(* Logix 5000 project; controller Almacen_2 vendor 1 type 14 code 235 rev 36.11; software revision 36.00; part 2 of 2 *)
(* tags used below, declared in another part *)
   Contador_Salida_Conveyor : COUNTER;
   End_Conveyor_Rutine : BOOL;
   PosDer_Alm_5_C : BOOL;
   PosDer_Alm_5_E : BOOL;
   PosIzq_Alm_7_C : BOOL;
   PosIzq_Conv_7_C : BOOL;
   PosIzq_Conv_8_C : BOOL;
   Recuperar_Pieza : BOOL;
   Recuperar_Pieza_Desde_RutinaConveyor : BOOL;
   Reset_RutinaFinal : BOOL;
   Start_Conveyor : BOOL;
   Start_Rutine_Conveyor_2 : BOOL;
   Stop_Conveyor_2 : BOOL;
   tag_switch : BOOL;
   tag_switch2 : BOOL;
   tag_switch3 : BOOL;
   Tag_switch4 : BOOL;
   tag_switch5 : BOOL;
   tag_switch6 : BOOL;
   tag_switch7 : BOOL;
   tag_switch8 : BOOL;
   tag_switch_almacen10 : BOOL;
   tag_switch_almacen11 : BOOL;
   tag_switch_almacen12 : BOOL;
   tag_switch_almacen13 : BOOL;
   tag_switch_almacen14 : BOOL;
   tag_switch_almacen15 : BOOL;
   tag_switch_almacen16 : BOOL;
   tag_switch_almacen17 : BOOL;
   tag_switch_almacen_abrir_gripper2 : BOOL;
   tag_switch_almacen_cerrar_gripper2 : BOOL;
   tag_timer_piston : BOOL;
   tag_timer_piston2 : BOOL;
   Timer10_Recuperar_Pieza : TIMER;
   Timer11_Posicion_Recuperar_Pieza : TIMER;
   Timer1_Cambio_Direccion_CNC : TIMER;
   Timer2 : TIMER;
   Timer3_Piston_Marcadora_OFF : TIMER;
   Timer4_Piston_Camara_ON : TIMER;
   Timer5_Piston_Camara_OFF : TIMER;
   Timer6_Cambio_Direccion_Almacen : TIMER;
   Timer7_Sensor_Entrada_Salida : TIMER;
   Timer8_End_RutinaConveyor : TIMER;
   Timer9_Piston_Salida : TIMER;
   Timer_Almacen_Abrir_Gripper2 : TIMER;
   Timer_Almacen_Cerrar_Gripper2 : TIMER;
   Timer_Almacen_Entrar_Posicion1_Regreso : TIMER;
   Timer_Almacen_Posicion_1_Regreso : TIMER;
   Timer_Almacen_Posicion_Above_Conveyor3 : TIMER;
   Timer_Almacen_Posicion_Above_Conveyor4 : TIMER;
   Timer_Almacen_Posicion_Conveyor2 : TIMER;
   Timer_Almacen_Posicion_Home3 : TIMER;
   Timer_Almacen_Posicion_Home4 : TIMER;
   Timer_Almacen_Salir_Posicion1_Regreso : TIMER;
   Estops_Ok : BOOL;
   Interlocks_Ok : BOOL;
   LigthCurtain2_Ok : BOOL;
   Run_Program_Almacen2 : BOOL;
   Safety_FromTEC81 : Safety;
   Sfty_OK : BOOL;
   Start_Almacen2 : BOOL;
   Start_Conveyor_2_From_RutinaFinal : BOOL;
   Start_Motor_Alm_2 : BOOL;
   Start_RutinaFinal : BOOL;
   tag_switch_almacen1 : BOOL;
   tag_switch_almacen2 : BOOL;
   tag_switch_almacen3 : BOOL;
   tag_switch_almacen4 : BOOL;
   tag_switch_almacen5 : BOOL;
   tag_switch_almacen6 : BOOL;
   tag_switch_almacen7 : BOOL;
   tag_switch_almacen8 : BOOL;
   tag_switch_almacen9 : BOOL;
   tag_switch_almacen_abrir_gripper : BOOL;
   tag_switch_almacen_cerrar_gripper : BOOL;
   Timer_Almacen_Abrir_Gripper : TIMER;
   Timer_Almacen_Cerrar_Gripper : TIMER;
   Timer_Almacen_Entrar_Posicion1 : TIMER;
   Timer_Almacen_Posicion1 : TIMER;
   Timer_Almacen_Posicion_Above_Conveyor : TIMER;
   Timer_Almacen_Posicion_Above_Conveyor2 : TIMER;
   Timer_Almacen_Posicion_Conveyor : TIMER;
   Timer_Almacen_Posicion_Giro_A_Conveyor : TIMER;
   Timer_Almacen_Posicion_Home : TIMER;
   Timer_Almacen_Posicion_Home2 : TIMER;
   Timer_Almacen_Salir_Posicion1 : TIMER;
(* MainProgram, continued *)

ROUTINE RutinaConveyor   (* ladder *)
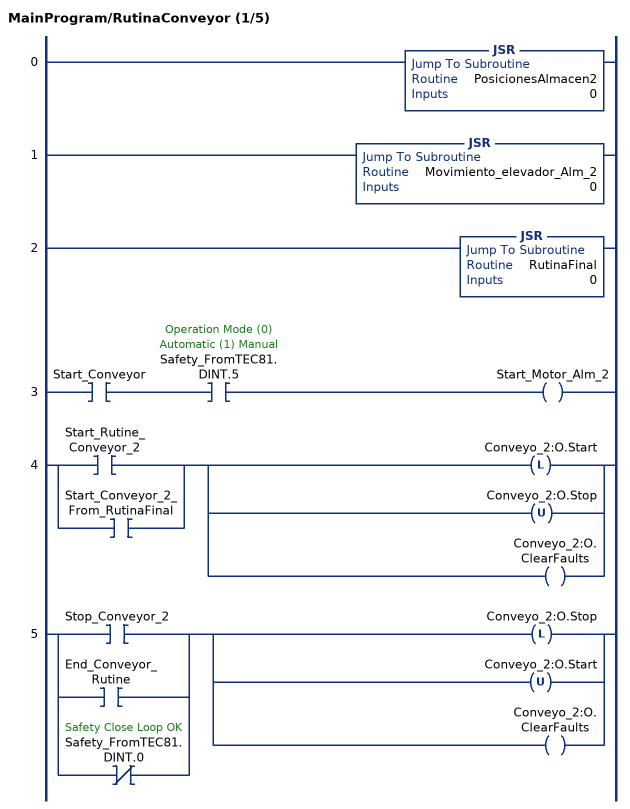
   0: JSR(PosicionesAlmacen2,0);
   1: JSR(Movimiento_elevador_Alm_2,0);
   2: JSR(RutinaFinal,0);
   3: XIC(Start_Conveyor)XIC(Safety_FromTEC81.DINT.5)OTE(Start_Motor_Alm_2);
   4: [XIC(Start_Rutine_Conveyor_2) ,XIC(Start_Conveyor_2_From_RutinaFinal) ][OTL(Conveyo_2:O.Start) ,OTU(Conveyo_2:O.Stop) ,OTE(Conveyo_2:O.ClearFaults) ];
   5: [XIC(Stop_Conveyor_2) ,XIC(End_Conveyor_Rutine) ,XIO(Safety_FromTEC81.DINT.0) ][OTL(Conveyo_2:O.Stop) ,OTU(Conveyo_2:O.Start) ,OTE(Conveyo_2:O.ClearFaults) ];
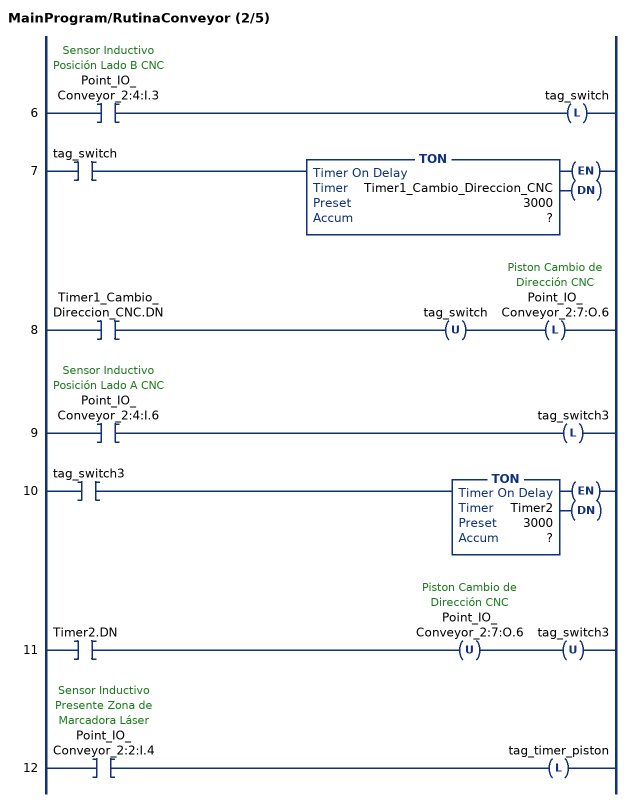
   6: XIC(Point_IO_Conveyor_2:4:I.3)OTL(tag_switch);
   7: XIC(tag_switch)TON(Timer1_Cambio_Direccion_CNC,?,?);
   8: XIC(Timer1_Cambio_Direccion_CNC.DN)OTU(tag_switch)OTL(Point_IO_Conveyor_2:7:O.6);
   9: XIC(Point_IO_Conveyor_2:4:I.6)OTL(tag_switch3);
   10: XIC(tag_switch3)TON(Timer2,?,?);
   11: XIC(Timer2.DN)OTU(Point_IO_Conveyor_2:7:O.6)OTU(tag_switch3);
   12: XIC(Point_IO_Conveyor_2:2:I.4)OTL(tag_timer_piston);
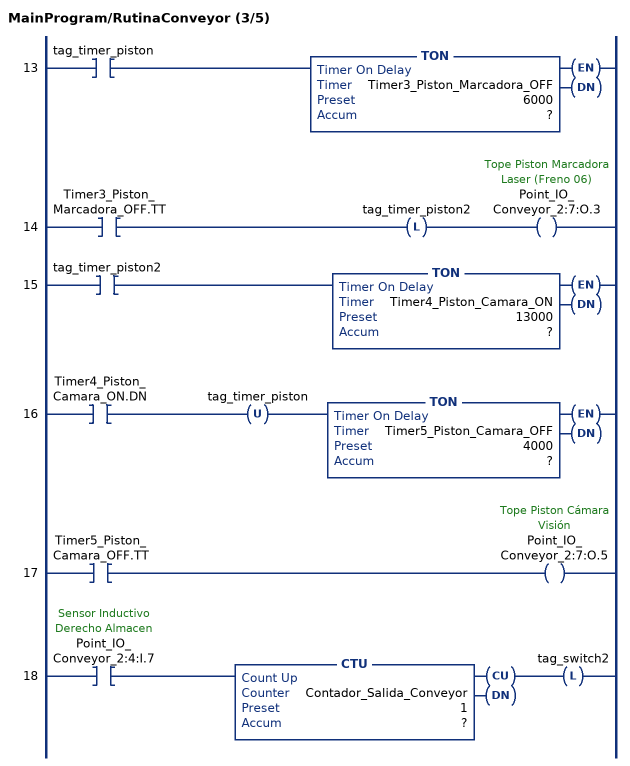
   13: XIC(tag_timer_piston)TON(Timer3_Piston_Marcadora_OFF,?,?);
   14: XIC(Timer3_Piston_Marcadora_OFF.TT)OTL(tag_timer_piston2)OTE(Point_IO_Conveyor_2:7:O.3);
   15: XIC(tag_timer_piston2)TON(Timer4_Piston_Camara_ON,?,?);
   16: XIC(Timer4_Piston_Camara_ON.DN)OTU(tag_timer_piston)TON(Timer5_Piston_Camara_OFF,?,?);
   17: XIC(Timer5_Piston_Camara_OFF.TT)OTE(Point_IO_Conveyor_2:7:O.5);
   18: XIC(Point_IO_Conveyor_2:4:I.7)CTU(Contador_Salida_Conveyor,?,?)OTL(tag_switch2);
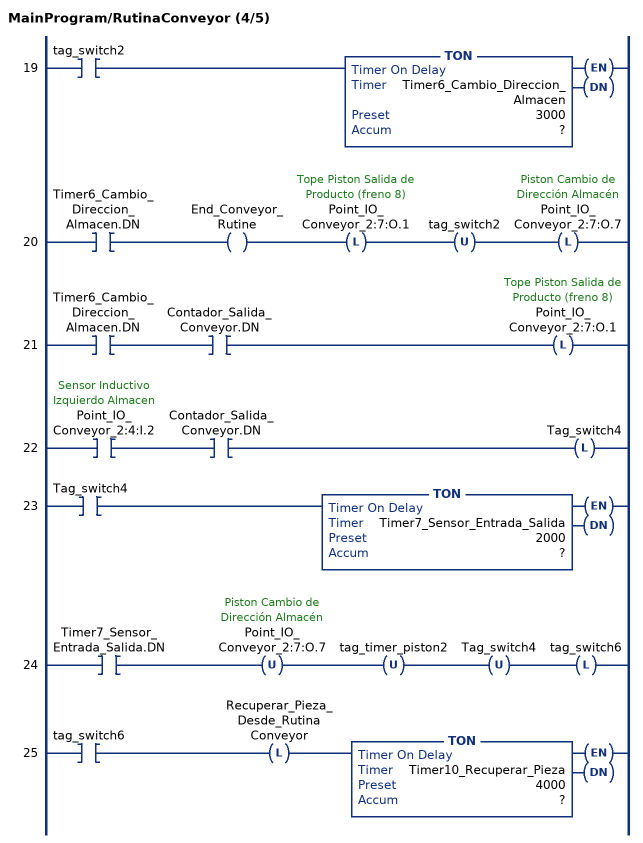
   19: XIC(tag_switch2)TON(Timer6_Cambio_Direccion_Almacen,?,?);
   20: XIC(Timer6_Cambio_Direccion_Almacen.DN)OTE(End_Conveyor_Rutine)OTL(Point_IO_Conveyor_2:7:O.1)OTU(tag_switch2)OTL(Point_IO_Conveyor_2:7:O.7);
   21: XIC(Timer6_Cambio_Direccion_Almacen.DN)XIC(Contador_Salida_Conveyor.DN)OTL(Point_IO_Conveyor_2:7:O.1);
   22: XIC(Point_IO_Conveyor_2:4:I.2)XIC(Contador_Salida_Conveyor.DN)OTL(Tag_switch4);
   23: XIC(Tag_switch4)TON(Timer7_Sensor_Entrada_Salida,?,?);
   24: XIC(Timer7_Sensor_Entrada_Salida.DN)OTU(Point_IO_Conveyor_2:7:O.7)OTU(tag_timer_piston2)OTU(Tag_switch4)OTL(tag_switch6);
   25: XIC(tag_switch6)OTL(Recuperar_Pieza_Desde_RutinaConveyor)TON(Timer10_Recuperar_Pieza,?,?);
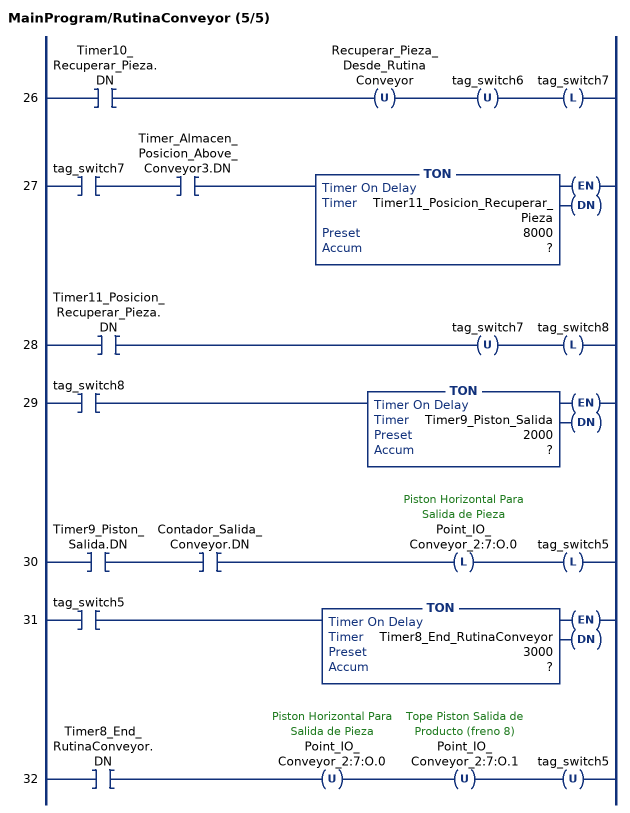
   26: XIC(Timer10_Recuperar_Pieza.DN)OTU(Recuperar_Pieza_Desde_RutinaConveyor)OTU(tag_switch6)OTL(tag_switch7);
   27: XIC(tag_switch7)XIC(Timer_Almacen_Posicion_Above_Conveyor3.DN)TON(Timer11_Posicion_Recuperar_Pieza,?,?);
   28: XIC(Timer11_Posicion_Recuperar_Pieza.DN)OTU(tag_switch7)OTL(tag_switch8);
   29: XIC(tag_switch8)TON(Timer9_Piston_Salida,?,?);
   30: XIC(Timer9_Piston_Salida.DN)XIC(Contador_Salida_Conveyor.DN)OTL(Point_IO_Conveyor_2:7:O.0)OTL(tag_switch5);
   31: XIC(tag_switch5)TON(Timer8_End_RutinaConveyor,?,?);
   32: XIC(Timer8_End_RutinaConveyor.DN)OTU(Point_IO_Conveyor_2:7:O.0)OTU(Point_IO_Conveyor_2:7:O.1)OTU(tag_switch5);
END_ROUTINE

ROUTINE RutinaFinal   (* ladder *)
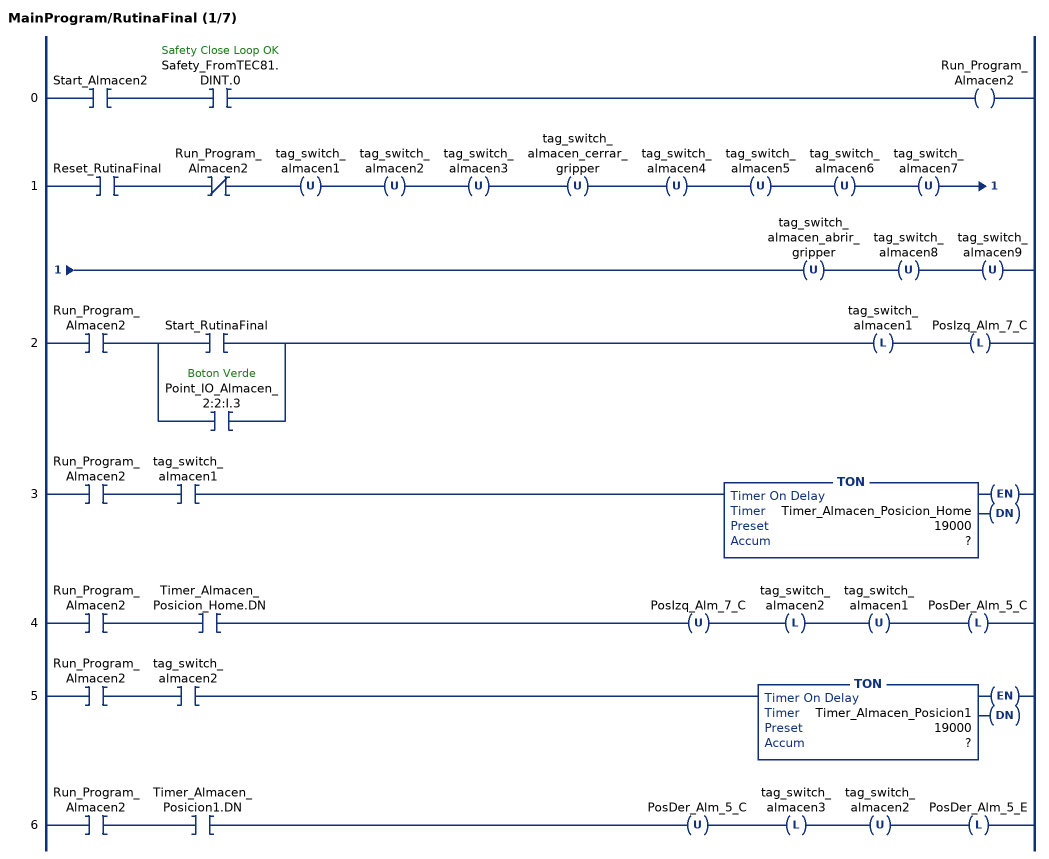
   0: XIC(Start_Almacen2)XIC(Safety_FromTEC81.DINT.0)OTE(Run_Program_Almacen2);
   1: XIC(Reset_RutinaFinal)XIO(Run_Program_Almacen2)OTU(tag_switch_almacen1)OTU(tag_switch_almacen2)OTU(tag_switch_almacen3)OTU(tag_switch_almacen_cerrar_gripper)OTU(tag_switch_almacen4)OTU(tag_switch_almacen5)OTU(tag_switch_almacen6)OTU(tag_switch_almacen7)OTU(tag_switch_almacen_abrir_gripper)OTU(tag_switch_almacen8)OTU(tag_switch_almacen9);
   2: XIC(Run_Program_Almacen2)[XIC(Start_RutinaFinal) ,XIC(Point_IO_Almacen_2:2:I.3) ]OTL(tag_switch_almacen1)OTL(PosIzq_Alm_7_C);
   3: XIC(Run_Program_Almacen2)XIC(tag_switch_almacen1)TON(Timer_Almacen_Posicion_Home,?,?);
   4: XIC(Run_Program_Almacen2)XIC(Timer_Almacen_Posicion_Home.DN)OTU(PosIzq_Alm_7_C)OTL(tag_switch_almacen2)OTU(tag_switch_almacen1)OTL(PosDer_Alm_5_C);
   5: XIC(Run_Program_Almacen2)XIC(tag_switch_almacen2)TON(Timer_Almacen_Posicion1,?,?);
   6: XIC(Run_Program_Almacen2)XIC(Timer_Almacen_Posicion1.DN)OTU(PosDer_Alm_5_C)OTL(tag_switch_almacen3)OTU(tag_switch_almacen2)OTL(PosDer_Alm_5_E);
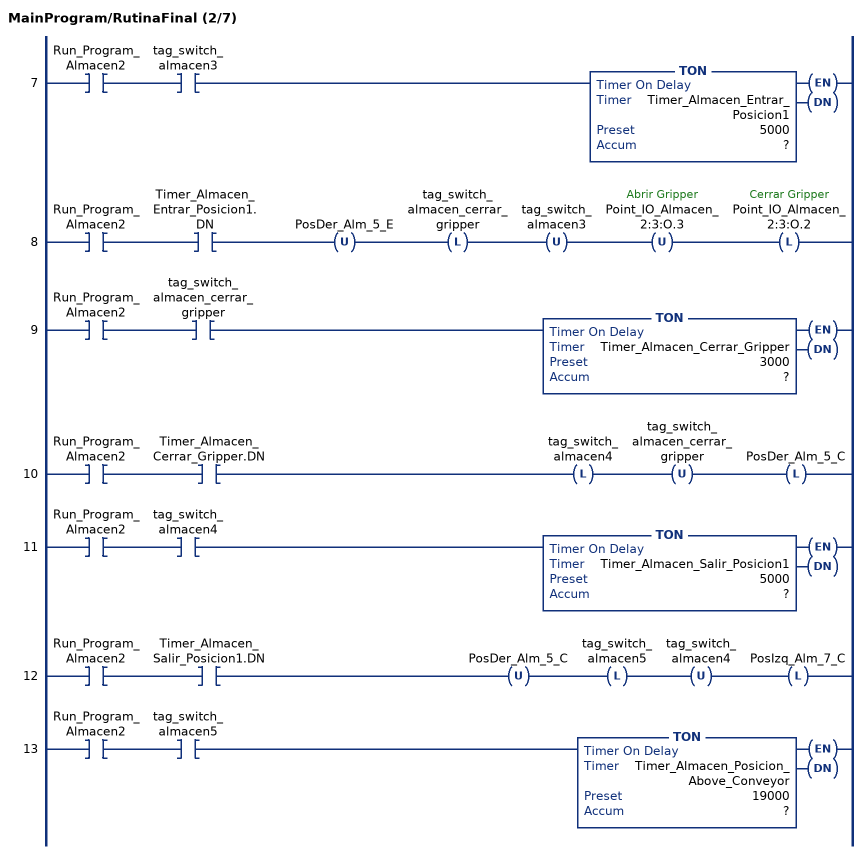
   7: XIC(Run_Program_Almacen2)XIC(tag_switch_almacen3)TON(Timer_Almacen_Entrar_Posicion1,?,?);
   8: XIC(Run_Program_Almacen2)XIC(Timer_Almacen_Entrar_Posicion1.DN)OTU(PosDer_Alm_5_E)OTL(tag_switch_almacen_cerrar_gripper)OTU(tag_switch_almacen3)OTU(Point_IO_Almacen_2:3:O.3)OTL(Point_IO_Almacen_2:3:O.2);
   9: XIC(Run_Program_Almacen2)XIC(tag_switch_almacen_cerrar_gripper)TON(Timer_Almacen_Cerrar_Gripper,?,?);
   10: XIC(Run_Program_Almacen2)XIC(Timer_Almacen_Cerrar_Gripper.DN)OTL(tag_switch_almacen4)OTU(tag_switch_almacen_cerrar_gripper)OTL(PosDer_Alm_5_C);
   11: XIC(Run_Program_Almacen2)XIC(tag_switch_almacen4)TON(Timer_Almacen_Salir_Posicion1,?,?);
   12: XIC(Run_Program_Almacen2)XIC(Timer_Almacen_Salir_Posicion1.DN)OTU(PosDer_Alm_5_C)OTL(tag_switch_almacen5)OTU(tag_switch_almacen4)OTL(PosIzq_Alm_7_C);
   13: XIC(Run_Program_Almacen2)XIC(tag_switch_almacen5)TON(Timer_Almacen_Posicion_Above_Conveyor,?,?);
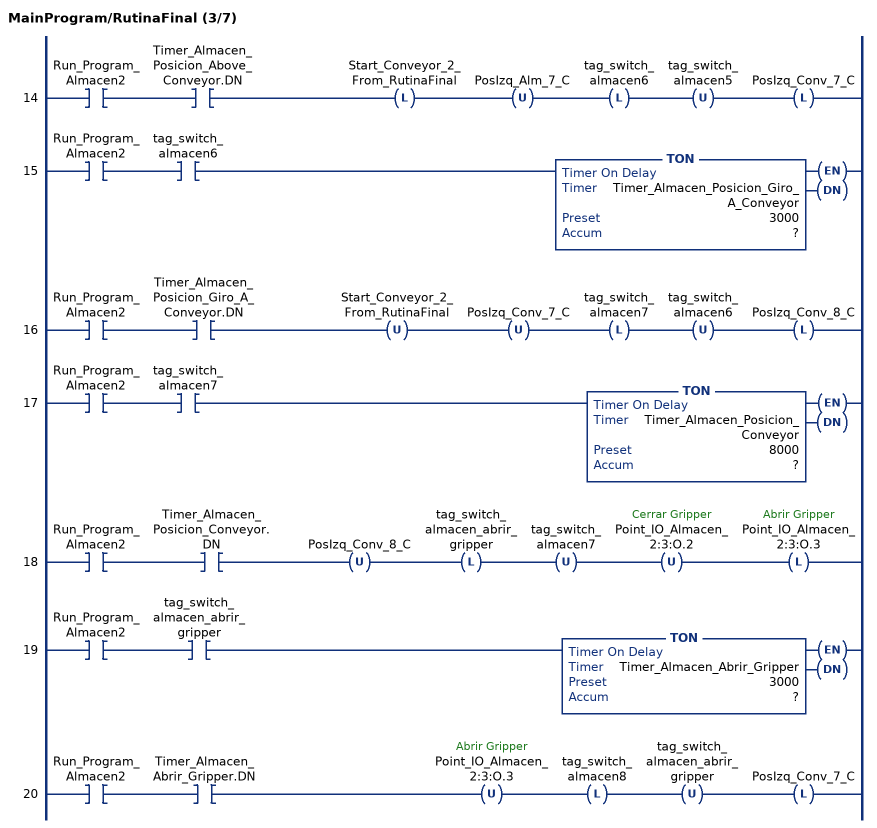
   14: XIC(Run_Program_Almacen2)XIC(Timer_Almacen_Posicion_Above_Conveyor.DN)OTL(Start_Conveyor_2_From_RutinaFinal)OTU(PosIzq_Alm_7_C)OTL(tag_switch_almacen6)OTU(tag_switch_almacen5)OTL(PosIzq_Conv_7_C);
   15: XIC(Run_Program_Almacen2)XIC(tag_switch_almacen6)TON(Timer_Almacen_Posicion_Giro_A_Conveyor,?,?);
   16: XIC(Run_Program_Almacen2)XIC(Timer_Almacen_Posicion_Giro_A_Conveyor.DN)OTU(Start_Conveyor_2_From_RutinaFinal)OTU(PosIzq_Conv_7_C)OTL(tag_switch_almacen7)OTU(tag_switch_almacen6)OTL(PosIzq_Conv_8_C);
   17: XIC(Run_Program_Almacen2)XIC(tag_switch_almacen7)TON(Timer_Almacen_Posicion_Conveyor,?,?);
   18: XIC(Run_Program_Almacen2)XIC(Timer_Almacen_Posicion_Conveyor.DN)OTU(PosIzq_Conv_8_C)OTL(tag_switch_almacen_abrir_gripper)OTU(tag_switch_almacen7)OTU(Point_IO_Almacen_2:3:O.2)OTL(Point_IO_Almacen_2:3:O.3);
   19: XIC(Run_Program_Almacen2)XIC(tag_switch_almacen_abrir_gripper)TON(Timer_Almacen_Abrir_Gripper,?,?);
   20: XIC(Run_Program_Almacen2)XIC(Timer_Almacen_Abrir_Gripper.DN)OTU(Point_IO_Almacen_2:3:O.3)OTL(tag_switch_almacen8)OTU(tag_switch_almacen_abrir_gripper)OTL(PosIzq_Conv_7_C);
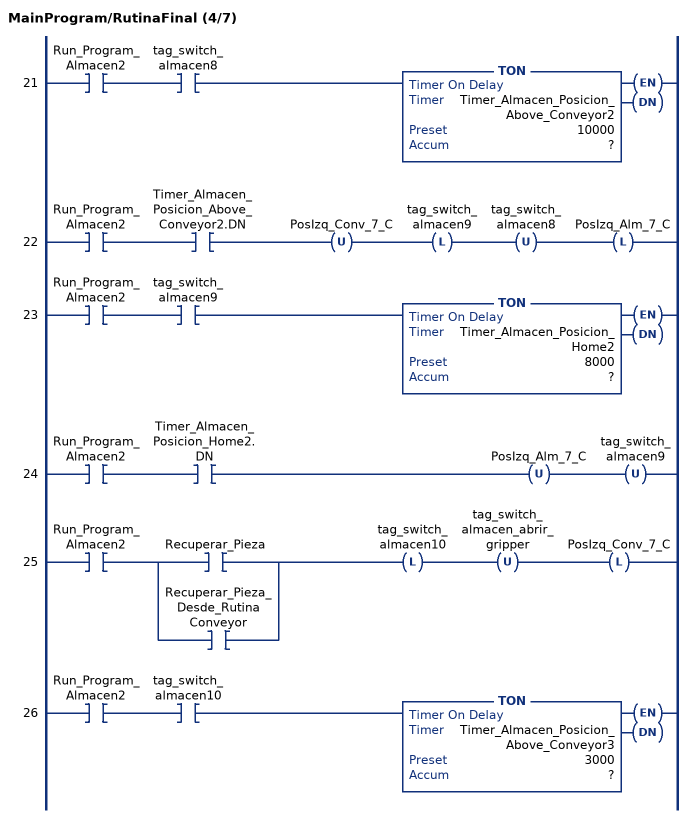
   21: XIC(Run_Program_Almacen2)XIC(tag_switch_almacen8)TON(Timer_Almacen_Posicion_Above_Conveyor2,?,?);
   22: XIC(Run_Program_Almacen2)XIC(Timer_Almacen_Posicion_Above_Conveyor2.DN)OTU(PosIzq_Conv_7_C)OTL(tag_switch_almacen9)OTU(tag_switch_almacen8)OTL(PosIzq_Alm_7_C);
   23: XIC(Run_Program_Almacen2)XIC(tag_switch_almacen9)TON(Timer_Almacen_Posicion_Home2,?,?);
   24: XIC(Run_Program_Almacen2)XIC(Timer_Almacen_Posicion_Home2.DN)OTU(PosIzq_Alm_7_C)OTU(tag_switch_almacen9);
   25: XIC(Run_Program_Almacen2)[XIC(Recuperar_Pieza) ,XIC(Recuperar_Pieza_Desde_RutinaConveyor) ]OTL(tag_switch_almacen10)OTU(tag_switch_almacen_abrir_gripper)OTL(PosIzq_Conv_7_C);
   26: XIC(Run_Program_Almacen2)XIC(tag_switch_almacen10)TON(Timer_Almacen_Posicion_Above_Conveyor3,?,?);
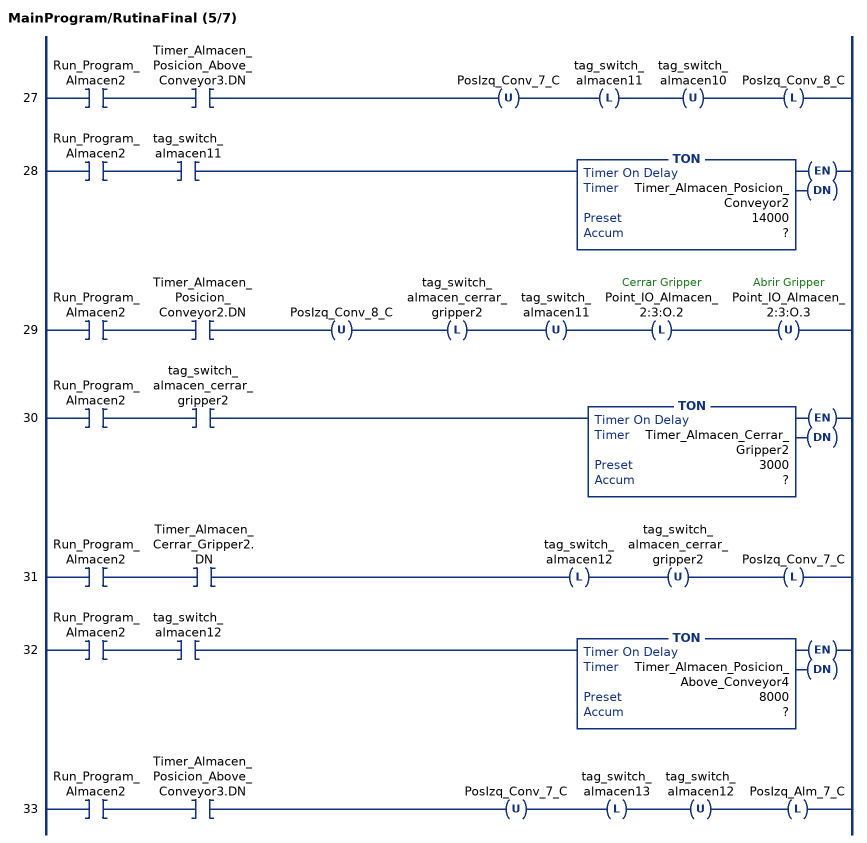
   27: XIC(Run_Program_Almacen2)XIC(Timer_Almacen_Posicion_Above_Conveyor3.DN)OTU(PosIzq_Conv_7_C)OTL(tag_switch_almacen11)OTU(tag_switch_almacen10)OTL(PosIzq_Conv_8_C);
   28: XIC(Run_Program_Almacen2)XIC(tag_switch_almacen11)TON(Timer_Almacen_Posicion_Conveyor2,?,?);
   29: XIC(Run_Program_Almacen2)XIC(Timer_Almacen_Posicion_Conveyor2.DN)OTU(PosIzq_Conv_8_C)OTL(tag_switch_almacen_cerrar_gripper2)OTU(tag_switch_almacen11)OTL(Point_IO_Almacen_2:3:O.2)OTU(Point_IO_Almacen_2:3:O.3);
   30: XIC(Run_Program_Almacen2)XIC(tag_switch_almacen_cerrar_gripper2)TON(Timer_Almacen_Cerrar_Gripper2,?,?);
   31: XIC(Run_Program_Almacen2)XIC(Timer_Almacen_Cerrar_Gripper2.DN)OTL(tag_switch_almacen12)OTU(tag_switch_almacen_cerrar_gripper2)OTL(PosIzq_Conv_7_C);
   32: XIC(Run_Program_Almacen2)XIC(tag_switch_almacen12)TON(Timer_Almacen_Posicion_Above_Conveyor4,?,?);
   33: XIC(Run_Program_Almacen2)XIC(Timer_Almacen_Posicion_Above_Conveyor3.DN)OTU(PosIzq_Conv_7_C)OTL(tag_switch_almacen13)OTU(tag_switch_almacen12)OTL(PosIzq_Alm_7_C);
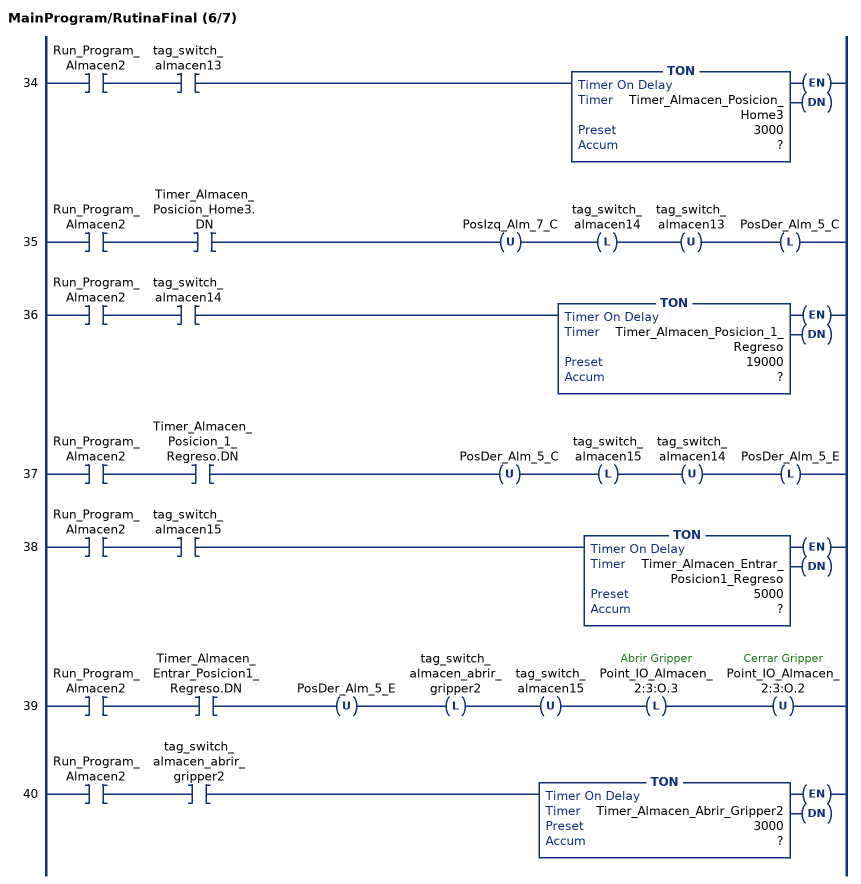
   34: XIC(Run_Program_Almacen2)XIC(tag_switch_almacen13)TON(Timer_Almacen_Posicion_Home3,?,?);
   35: XIC(Run_Program_Almacen2)XIC(Timer_Almacen_Posicion_Home3.DN)OTU(PosIzq_Alm_7_C)OTL(tag_switch_almacen14)OTU(tag_switch_almacen13)OTL(PosDer_Alm_5_C);
   36: XIC(Run_Program_Almacen2)XIC(tag_switch_almacen14)TON(Timer_Almacen_Posicion_1_Regreso,?,?);
   37: XIC(Run_Program_Almacen2)XIC(Timer_Almacen_Posicion_1_Regreso.DN)OTU(PosDer_Alm_5_C)OTL(tag_switch_almacen15)OTU(tag_switch_almacen14)OTL(PosDer_Alm_5_E);
   38: XIC(Run_Program_Almacen2)XIC(tag_switch_almacen15)TON(Timer_Almacen_Entrar_Posicion1_Regreso,?,?);
   39: XIC(Run_Program_Almacen2)XIC(Timer_Almacen_Entrar_Posicion1_Regreso.DN)OTU(PosDer_Alm_5_E)OTL(tag_switch_almacen_abrir_gripper2)OTU(tag_switch_almacen15)OTL(Point_IO_Almacen_2:3:O.3)OTU(Point_IO_Almacen_2:3:O.2);
   40: XIC(Run_Program_Almacen2)XIC(tag_switch_almacen_abrir_gripper2)TON(Timer_Almacen_Abrir_Gripper2,?,?);
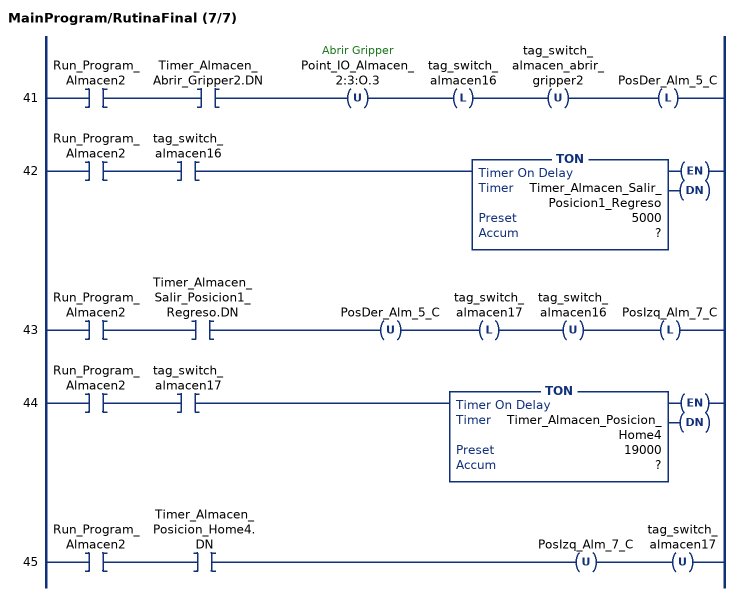
   41: XIC(Run_Program_Almacen2)XIC(Timer_Almacen_Abrir_Gripper2.DN)OTU(Point_IO_Almacen_2:3:O.3)OTL(tag_switch_almacen16)OTU(tag_switch_almacen_abrir_gripper2)OTL(PosDer_Alm_5_C);
   42: XIC(Run_Program_Almacen2)XIC(tag_switch_almacen16)TON(Timer_Almacen_Salir_Posicion1_Regreso,?,?);
   43: XIC(Run_Program_Almacen2)XIC(Timer_Almacen_Salir_Posicion1_Regreso.DN)OTU(PosDer_Alm_5_C)OTL(tag_switch_almacen17)OTU(tag_switch_almacen16)OTL(PosIzq_Alm_7_C);
   44: XIC(Run_Program_Almacen2)XIC(tag_switch_almacen17)TON(Timer_Almacen_Posicion_Home4,?,?);
   45: XIC(Run_Program_Almacen2)XIC(Timer_Almacen_Posicion_Home4.DN)OTU(PosIzq_Alm_7_C)OTU(tag_switch_almacen17);
END_ROUTINE
END_PROGRAM

PROGRAM SafetyProgram   (* main routine MainRoutine, safety *)

ROUTINE External_COMM   (* ladder *)
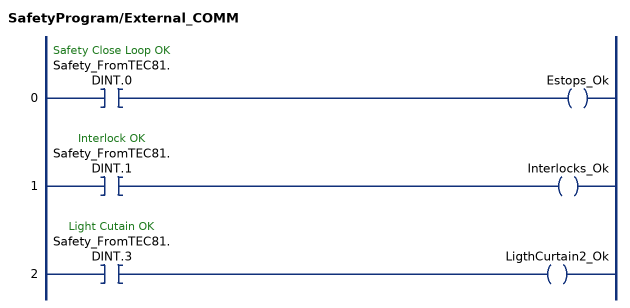
   0: XIC(Safety_FromTEC81.DINT.0)OTE(Estops_Ok);
   1: XIC(Safety_FromTEC81.DINT.1)OTE(Interlocks_Ok);
   2: XIC(Safety_FromTEC81.DINT.3)OTE(LigthCurtain2_Ok);
END_ROUTINE

ROUTINE MainRoutine   (* ladder *)
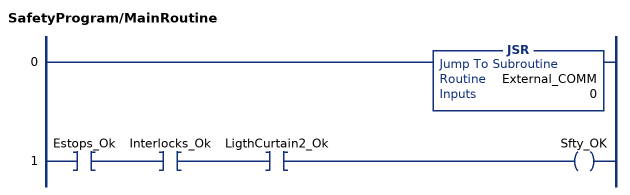
   0: JSR(External_COMM,0);
   1: XIC(Estops_Ok)XIC(Interlocks_Ok)XIC(LigthCurtain2_Ok)OTE(Sfty_OK);
END_ROUTINE
END_PROGRAM
